   "Carrier_37_SpareSafetyOutput(3_4)" AT %I2215.4 : Bool;   // SPARE SAFETY OUTPUT
   "Carrier_37_SpareSafetyOutput(3_5)" AT %I2215.5 : Bool;   // SPARE SAFETY OUTPUT
   "Carrier_37_SpareSafetyOutput(3_6)" AT %I2215.6 : Bool;   // SPARE SAFETY OUTPUT
   "Carrier_37_SpareSafetyOutput(3_7)" AT %I2215.7 : Bool;   // SPARE SAFETY OUTPUT
   "Carrier_37_Slot4_Input" AT %IW2216 : Word;   // SLOT 4 INPUT WORD
   "Carrier_37_480VPowerOn_MDCB1" AT %I2216.0 : Bool;   // 480 VAC POWER ON MDCB 1
   "Carrier_37_SpareInput(4_1)" AT %I2216.1 : Bool;   // SPARE INPUT
   "Carrier_37_SpareInput(4_2)" AT %I2216.2 : Bool;   // SPARE INPUT
   "Carrier_37_SitopSelectStatus" AT %I2216.3 : Bool;   // SITOP SELECT STATUS
   "Carrier_37_DCsupplyOnPSCB2" AT %I2216.4 : Bool;   // DC SUPPLY ON PSCB 2
   "Carrier_37_SpareInput(4_5)" AT %I2216.5 : Bool;   // SPARE INPUT
   "Carrier_37_SpareInput(4_6)" AT %I2216.6 : Bool;   // SPARE INPUT
   "Carrier_37_SpareInput(4_7)" AT %I2216.7 : Bool;   // SPARE INPUT
   "Carrier_37_PB1_ProdHoldLH" AT %I2217.0 : Bool;   // PB 1 PRODUCTION HOLD LH
   "Carrier_37_PB2_ResetLH" AT %I2217.1 : Bool;   // PB 2 RESET LH
   "Carrier_37_PB3_ProdHoldRH" AT %I2217.2 : Bool;   // PB 3 PRODUCTION HOLD RH
   "Carrier_37_PB4_ResetRH" AT %I2217.3 : Bool;   // PB 4 RESET RH
   "Carrier_37_SpareInput(4_14)" AT %I2217.4 : Bool;   // SPARE INPUT
   "Carrier_37_SpareInput(4_15)" AT %I2217.5 : Bool;   // SPARE INPUT
   "Carrier_37_SpareInput(4_16)" AT %I2217.6 : Bool;   // SPARE INPUT
   "Carrier_37_SpareInput(4_17)" AT %I2217.7 : Bool;   // SPARE INPUT
   "Carrier_37_Slot5_Output" AT %IW2218 : Word;   // SLOT 5 OUTPUT WORD
   "Carrier_37_IRD400_HMI_24VDC_ENABLE" AT %I2218.0 : Bool;   // IRD 400 PANEL HMI 24V DC POWER
   "Carrier_37_FaultLight_LH" AT %I2218.1 : Bool;   // FAULT LIGHT LH
   "Carrier_37_RunLight_LH" AT %I2218.2 : Bool;   // RUN LIGHT LH
   "Carrier_37_FaultLight_RH" AT %I2218.3 : Bool;   // FAULT LIGHT RH
   "Carrier_37_RunLight_RH" AT %I2218.4 : Bool;   // RUN LIGHT RH
   "Carrier_37_SpareOutput(5_5)" AT %I2218.5 : Bool;   // SPARE OUTPUT
   "Carrier_37_SpareOutput(5_6)" AT %I2218.6 : Bool;   // SPARE OUTPUT
   "Carrier_37_SpareOutput(5_7)" AT %I2218.7 : Bool;   // SPARE OUTPUT
   "Carrier_37_ActualSpeed" AT %IW2220 : Word;   // ACTUAL SPEED
   "Carrier_37_CarrierDriveAlarm" AT %IW2222 : Word;   // CARRIER DRIVE ALARM
   "Carrier_37_CarrierDriveWarning" AT %IW2224 : Word;   // CARRIER DRIVE WARNING
   "Carrier_38_Status" AT %IW2250 : Word;   // CARRIER STATUS WORD
   "Carrier_38_Status.0" AT %I2250.0 : Bool;   // HEARTBEAT
   "Carrier_38_Status.1" AT %I2250.1 : Bool;   // MANUAL
   "Carrier_38_Status.2" AT %I2250.2 : Bool;   // IN_AUTO
   "Carrier_38_Status.3" AT %I2250.3 : Bool;   // POSITIONING_COMPLETE
   "Carrier_38_Status.4" AT %I2250.4 : Bool;   // PRODUCTION HOLD
   "Carrier_38_Status.5" AT %I2250.5 : Bool;   // CARRIER MOVING FORWARD
   "Carrier_38_Status.6" AT %I2250.6 : Bool;   // CARRIER MOVING REVERSE
   "Carrier_38_Status.7" AT %I2250.7 : Bool;   // CARRIER FAULT
   "Carrier_38_Status.8" AT %I2251.0 : Bool;   // CRASH DETECT TRIPPED
   "Carrier_38_Status.9" AT %I2251.1 : Bool;
   "Carrier_38_Status.10" AT %I2251.2 : Bool;
   "Carrier_38_Status.11" AT %I2251.3 : Bool;
   "Carrier_38_Status.12" AT %I2251.4 : Bool;
   "Carrier_38_Status.13" AT %I2251.5 : Bool;
   "Carrier_38_Status.14" AT %I2251.6 : Bool;
   "Carrier_38_Status.15" AT %I2251.7 : Bool;
   "Carrier_38_SDCFaultCode" AT %IW2252 : Word;   // SDC FAULT CODE
   "Carrier_38_CarrierPosition" AT %ID2254 : DWord;   // CARRIER POSITION
   "Carrier_38_CarrierNumber" AT %IW2258 : Word;   // CARRIER NUMBER
   "Carrier_38_G120DControlWord" AT %IW2260 : Word;   // G120D_STW1_CONTROL
   "Carrier_38_G120DControlWord.0" AT %I2260.0 : Bool;   // Bit_00_ON
   "Carrier_38_G120DControlWord.1" AT %I2260.1 : Bool;   // Bit_01_AUS2_INH
   "Carrier_38_G120DControlWord.2" AT %I2260.2 : Bool;   // Bit_02_AUS3_STOP
   "Carrier_38_G120DControlWord.3" AT %I2260.3 : Bool;   // Bit_03_EN
   "Carrier_38_G120DControlWord.4" AT %I2260.4 : Bool;   // Bit_04_EN_RAMP
   "Carrier_38_G120DControlWord.5" AT %I2260.5 : Bool;   // Bit_05_START_RAMP
   "Carrier_38_G120DControlWord.6" AT %I2260.6 : Bool;   // Bit_06_SETPOINT
   "Carrier_38_G120DControlWord.7" AT %I2260.7 : Bool;   // Bit_07_RESET
   "Carrier_38_G120DControlWord.8" AT %I2261.0 : Bool;   // Bit_08_JOG_R
   "Carrier_38_G120DControlWord.9" AT %I2261.1 : Bool;   // Bit_09_JOG_L
   "Carrier_38_G120DControlWord.10" AT %I2261.2 : Bool;   // Bit_10_CONTR_PLC
   "Carrier_38_G120DControlWord.11" AT %I2261.3 : Bool;   // Bit_11_REVERSE
   "Carrier_38_G120DControlWord.12" AT %I2261.4 : Bool;   // Bit_12_BRAKE_RELEASE
   "Carrier_38_G120DControlWord.13" AT %I2261.5 : Bool;   // Bit_13_DDS
   "Carrier_38_G120DControlWord.14" AT %I2261.6 : Bool;   // Bit_14_DO0
   "Carrier_38_G120DControlWord.15" AT %I2261.7 : Bool;   // Bit_15_DO1
   "Carrier_38_G120DStatusWord" AT %IW2262 : Word;   // G120D_ZSW1_STATUS
   "Carrier_38_G120DStatusWord.0" AT %I2262.0 : Bool;   // Bit_00_READY_RUN
   "Carrier_38_G120DStatusWord.1" AT %I2262.1 : Bool;   // Bit_01_READY_ON
   "Carrier_38_G120DStatusWord.2" AT %I2262.2 : Bool;   // Bit_02_ENABLE
   "Carrier_38_G120DStatusWord.3" AT %I2262.3 : Bool;   // Bit_03_FAULT
   "Carrier_38_G120DStatusWord.4" AT %I2262.4 : Bool;   // Bit_04_OFF2
   "Carrier_38_G120DStatusWord.5" AT %I2262.5 : Bool;   // Bit_05_OFF3
   "Carrier_38_G120DStatusWord.6" AT %I2262.6 : Bool;   // Bit_06_LOCK_OUT
   "Carrier_38_G120DStatusWord.7" AT %I2262.7 : Bool;   // Bit_07_WARN
   "Carrier_38_G120DStatusWord.8" AT %I2263.0 : Bool;   // Bit_08_NO_DEVIATION
   "Carrier_38_G120DStatusWord.9" AT %I2263.1 : Bool;   // Bit_09_CONTR_PLC
   "Carrier_38_G120DStatusWord.10" AT %I2263.2 : Bool;   // Bit_10_F_MAX
   "Carrier_38_G120DStatusWord.11" AT %I2263.3 : Bool;   // Bit_11_LIMIT_REACHED
   "Carrier_38_G120DStatusWord.12" AT %I2263.4 : Bool;   // Bit_12_BRAKE_OPEN
   "Carrier_38_G120DStatusWord.13" AT %I2263.5 : Bool;   // Bit_13_NO_OVERTEMP
   "Carrier_38_G120DStatusWord.14" AT %I2263.6 : Bool;   // Bit_14_CW_CCW
   "Carrier_38_G120DStatusWord.15" AT %I2263.7 : Bool;   // Bit_15_OVERL
   "Carrier_38_Slot2_Input" AT %IW2264 : Word;   // SLOT 2 INPUT WORD
   "Carrier_38_CrashDetectSW" AT %I2264.0 : Bool;   // CRASH DETECT SW
   "Carrier_38_SpareSafetyInput(2_1)" AT %I2264.1 : Bool;   // SPARE SAFETY INPUT
   "Carrier_38_SpareSafetyInput(2_2)" AT %I2264.2 : Bool;   // SPARE SAFETY INPUT
   "Carrier_38_SpareSafetyInput(2_3)" AT %I2264.3 : Bool;   // SPARE SAFETY INPUT
   "Carrier_38_SpareSafetyInput(2_4)" AT %I2264.4 : Bool;   // SPARE SAFETY INPUT
   "Carrier_38_SpareSafetyInput(2_5)" AT %I2264.5 : Bool;   // SPARE SAFETY INPUT
   "Carrier_38_SpareSafetyInput(2_6)" AT %I2264.6 : Bool;   // SPARE SAFETY INPUT
   "Carrier_38_SpareSafetyInput(2_7)" AT %I2264.7 : Bool;   // SPARE SAFETY INPUT
   "Carrier_38_Slot3_SafetyOutput" AT %IW2265 : Word;   // SLOT 3 SAFETY OUTPUT WORD
   "Carrier_38_Crash_Detect_OK" AT %I2265.0 : Bool;   // CARRIER CRASH DETECT
   "Carrier_38_SpareSafetyOutput(3_1)" AT %I2265.1 : Bool;   // SPARE SAFETY OUTPUT
   "Carrier_38_SpareSafetyOutput(3_2)" AT %I2265.2 : Bool;   // SPARE SAFETY OUTPUT
   "Carrier_38_SpareSafetyOutput(3_3)" AT %I2265.3 : Bool;   // SPARE SAFETY OUTPUT
   "Carrier_38_SpareSafetyOutput(3_4)" AT %I2265.4 : Bool;   // SPARE SAFETY OUTPUT
   "Carrier_38_SpareSafetyOutput(3_5)" AT %I2265.5 : Bool;   // SPARE SAFETY OUTPUT
   "Carrier_38_SpareSafetyOutput(3_6)" AT %I2265.6 : Bool;   // SPARE SAFETY OUTPUT
   "Carrier_38_SpareSafetyOutput(3_7)" AT %I2265.7 : Bool;   // SPARE SAFETY OUTPUT
   "Carrier_38_Slot4_Input" AT %IW2266 : Word;   // SLOT 4 INPUT WORD
   "Carrier_38_480VPowerOn_MDCB1" AT %I2266.0 : Bool;   // 480 VAC POWER ON MDCB 1
   "Carrier_38_SpareInput(4_1)" AT %I2266.1 : Bool;   // SPARE INPUT
   "Carrier_38_SpareInput(4_2)" AT %I2266.2 : Bool;   // SPARE INPUT
   "Carrier_38_SitopSelectStatus" AT %I2266.3 : Bool;   // SITOP SELECT STATUS
   "Carrier_38_DCsupplyOnPSCB2" AT %I2266.4 : Bool;   // DC SUPPLY ON PSCB 2
   "Carrier_38_SpareInput(4_5)" AT %I2266.5 : Bool;   // SPARE INPUT
   "Carrier_38_SpareInput(4_6)" AT %I2266.6 : Bool;   // SPARE INPUT
   "Carrier_38_SpareInput(4_7)" AT %I2266.7 : Bool;   // SPARE INPUT
   "Carrier_38_PB1_ProdHoldLH" AT %I2267.0 : Bool;   // PB 1 PRODUCTION HOLD LH
   "Carrier_38_PB2_ResetLH" AT %I2267.1 : Bool;   // PB 2 RESET LH
   "Carrier_38_PB3_ProdHoldRH" AT %I2267.2 : Bool;   // PB 3 PRODUCTION HOLD RH
   "Carrier_38_PB4_ResetRH" AT %I2267.3 : Bool;   // PB 4 RESET RH
   "Carrier_38_SpareInput(4_14)" AT %I2267.4 : Bool;   // SPARE INPUT
   "Carrier_38_SpareInput(4_15)" AT %I2267.5 : Bool;   // SPARE INPUT
   "Carrier_38_SpareInput(4_16)" AT %I2267.6 : Bool;   // SPARE INPUT
   "Carrier_38_SpareInput(4_17)" AT %I2267.7 : Bool;   // SPARE INPUT
   "Carrier_38_Slot5_Output" AT %IW2268 : Word;   // SLOT 5 OUTPUT WORD
   "Carrier_38_IRD400_HMI_24VDC_ENABLE" AT %I2268.0 : Bool;   // IRD 400 PANEL HMI 24V DC POWER
   "Carrier_38_FaultLight_LH" AT %I2268.1 : Bool;   // FAULT LIGHT LH
   "Carrier_38_RunLight_LH" AT %I2268.2 : Bool;   // RUN LIGHT LH
   "Carrier_38_FaultLight_RH" AT %I2268.3 : Bool;   // FAULT LIGHT RH
   "Carrier_38_RunLight_RH" AT %I2268.4 : Bool;   // RUN LIGHT RH
   "Carrier_38_SpareOutput(5_5)" AT %I2268.5 : Bool;   // SPARE OUTPUT
   "Carrier_38_SpareOutput(5_6)" AT %I2268.6 : Bool;   // SPARE OUTPUT
   "Carrier_38_SpareOutput(5_7)" AT %I2268.7 : Bool;   // SPARE OUTPUT
   "Carrier_38_ActualSpeed" AT %IW2270 : Word;   // ACTUAL SPEED
   "Carrier_38_CarrierDriveAlarm" AT %IW2272 : Word;   // CARRIER DRIVE ALARM
   "Carrier_38_CarrierDriveWarning" AT %IW2274 : Word;   // CARRIER DRIVE WARNING
   "Carrier_39_Status" AT %IW2300 : Word;   // CARRIER STATUS WORD
   "Carrier_39_Status.0" AT %I2300.0 : Bool;   // HEARTBEAT
   "Carrier_39_Status.1" AT %I2300.1 : Bool;   // MANUAL
   "Carrier_39_Status.2" AT %I2300.2 : Bool;   // IN_AUTO
   "Carrier_39_Status.3" AT %I2300.3 : Bool;   // POSITIONING_COMPLETE
   "Carrier_39_Status.4" AT %I2300.4 : Bool;   // PRODUCTION HOLD
   "Carrier_39_Status.5" AT %I2300.5 : Bool;   // CARRIER MOVING FORWARD
   "Carrier_39_Status.6" AT %I2300.6 : Bool;   // CARRIER MOVING REVERSE
   "Carrier_39_Status.7" AT %I2300.7 : Bool;   // CARRIER FAULT
   "Carrier_39_Status.8" AT %I2301.0 : Bool;   // CRASH DETECT TRIPPED
   "Carrier_39_Status.9" AT %I2301.1 : Bool;
   "Carrier_39_Status.10" AT %I2301.2 : Bool;
   "Carrier_39_Status.11" AT %I2301.3 : Bool;
   "Carrier_39_Status.12" AT %I2301.4 : Bool;
   "Carrier_39_Status.13" AT %I2301.5 : Bool;
   "Carrier_39_Status.14" AT %I2301.6 : Bool;
   "Carrier_39_Status.15" AT %I2301.7 : Bool;
   "Carrier_39_SDCFaultCode" AT %IW2302 : Word;   // SDC FAULT CODE
   "Carrier_39_CarrierPosition" AT %ID2304 : DWord;   // CARRIER POSITION
   "Carrier_39_CarrierNumber" AT %IW2308 : Word;   // CARRIER NUMBER
   "Carrier_39_G120DControlWord" AT %IW2310 : Word;   // G120D_STW1_CONTROL
   "Carrier_39_G120DControlWord.0" AT %I2310.0 : Bool;   // Bit_00_ON
   "Carrier_39_G120DControlWord.1" AT %I2310.1 : Bool;   // Bit_01_AUS2_INH
   "Carrier_39_G120DControlWord.2" AT %I2310.2 : Bool;   // Bit_02_AUS3_STOP
   "Carrier_39_G120DControlWord.3" AT %I2310.3 : Bool;   // Bit_03_EN
   "Carrier_39_G120DControlWord.4" AT %I2310.4 : Bool;   // Bit_04_EN_RAMP
   "Carrier_39_G120DControlWord.5" AT %I2310.5 : Bool;   // Bit_05_START_RAMP
   "Carrier_39_G120DControlWord.6" AT %I2310.6 : Bool;   // Bit_06_SETPOINT
   "Carrier_39_G120DControlWord.7" AT %I2310.7 : Bool;   // Bit_07_RESET
   "Carrier_39_G120DControlWord.8" AT %I2311.0 : Bool;   // Bit_08_JOG_R
   "Carrier_39_G120DControlWord.9" AT %I2311.1 : Bool;   // Bit_09_JOG_L
   "Carrier_39_G120DControlWord.10" AT %I2311.2 : Bool;   // Bit_10_CONTR_PLC
   "Carrier_39_G120DControlWord.11" AT %I2311.3 : Bool;   // Bit_11_REVERSE
   "Carrier_39_G120DControlWord.12" AT %I2311.4 : Bool;   // Bit_12_BRAKE_RELEASE
   "Carrier_39_G120DControlWord.13" AT %I2311.5 : Bool;   // Bit_13_DDS
   "Carrier_39_G120DControlWord.14" AT %I2311.6 : Bool;   // Bit_14_DO0
   "Carrier_39_G120DControlWord.15" AT %I2311.7 : Bool;   // Bit_15_DO1
   "Carrier_39_G120DStatusWord" AT %IW2312 : Word;   // G120D_ZSW1_STATUS
   "Carrier_39_G120DStatusWord.0" AT %I2312.0 : Bool;   // Bit_00_READY_RUN
   "Carrier_39_G120DStatusWord.1" AT %I2312.1 : Bool;   // Bit_01_READY_ON
   "Carrier_39_G120DStatusWord.2" AT %I2312.2 : Bool;   // Bit_02_ENABLE
   "Carrier_39_G120DStatusWord.3" AT %I2312.3 : Bool;   // Bit_03_FAULT
   "Carrier_39_G120DStatusWord.4" AT %I2312.4 : Bool;   // Bit_04_OFF2
   "Carrier_39_G120DStatusWord.5" AT %I2312.5 : Bool;   // Bit_05_OFF3
   "Carrier_39_G120DStatusWord.6" AT %I2312.6 : Bool;   // Bit_06_LOCK_OUT
   "Carrier_39_G120DStatusWord.7" AT %I2312.7 : Bool;   // Bit_07_WARN
   "Carrier_39_G120DStatusWord.8" AT %I2313.0 : Bool;   // Bit_08_NO_DEVIATION
   "Carrier_39_G120DStatusWord.9" AT %I2313.1 : Bool;   // Bit_09_CONTR_PLC
   "Carrier_39_G120DStatusWord.10" AT %I2313.2 : Bool;   // Bit_10_F_MAX
   "Carrier_39_G120DStatusWord.11" AT %I2313.3 : Bool;   // Bit_11_LIMIT_REACHED
   "Carrier_39_G120DStatusWord.12" AT %I2313.4 : Bool;   // Bit_12_BRAKE_OPEN
   "Carrier_39_G120DStatusWord.13" AT %I2313.5 : Bool;   // Bit_13_NO_OVERTEMP
   "Carrier_39_G120DStatusWord.14" AT %I2313.6 : Bool;   // Bit_14_CW_CCW
   "Carrier_39_G120DStatusWord.15" AT %I2313.7 : Bool;   // Bit_15_OVERL
   "Carrier_39_Slot2_Input" AT %IW2314 : Word;   // SLOT 2 INPUT WORD
   "Carrier_39_CrashDetectSW" AT %I2314.0 : Bool;   // CRASH DETECT SW
   "Carrier_39_SpareSafetyInput(2_1)" AT %I2314.1 : Bool;   // SPARE SAFETY INPUT
   "Carrier_39_SpareSafetyInput(2_2)" AT %I2314.2 : Bool;   // SPARE SAFETY INPUT
   "Carrier_39_SpareSafetyInput(2_3)" AT %I2314.3 : Bool;   // SPARE SAFETY INPUT
   "Carrier_39_SpareSafetyInput(2_4)" AT %I2314.4 : Bool;   // SPARE SAFETY INPUT
   "Carrier_39_SpareSafetyInput(2_5)" AT %I2314.5 : Bool;   // SPARE SAFETY INPUT
   "Carrier_39_SpareSafetyInput(2_6)" AT %I2314.6 : Bool;   // SPARE SAFETY INPUT
   "Carrier_39_SpareSafetyInput(2_7)" AT %I2314.7 : Bool;   // SPARE SAFETY INPUT
   "Carrier_39_Slot3_SafetyOutput" AT %IW2315 : Word;   // SLOT 3 SAFETY OUTPUT WORD
   "Carrier_39_Crash_Detect_OK" AT %I2315.0 : Bool;   // CARRIER CRASH DETECT
   "Carrier_39_SpareSafetyOutput(3_1)" AT %I2315.1 : Bool;   // SPARE SAFETY OUTPUT
   "Carrier_39_SpareSafetyOutput(3_2)" AT %I2315.2 : Bool;   // SPARE SAFETY OUTPUT
   "Carrier_39_SpareSafetyOutput(3_3)" AT %I2315.3 : Bool;   // SPARE SAFETY OUTPUT
   "Carrier_39_SpareSafetyOutput(3_4)" AT %I2315.4 : Bool;   // SPARE SAFETY OUTPUT
   "Carrier_39_SpareSafetyOutput(3_5)" AT %I2315.5 : Bool;   // SPARE SAFETY OUTPUT
   "Carrier_39_SpareSafetyOutput(3_6)" AT %I2315.6 : Bool;   // SPARE SAFETY OUTPUT
   "Carrier_39_SpareSafetyOutput(3_7)" AT %I2315.7 : Bool;   // SPARE SAFETY OUTPUT
   "Carrier_39_Slot4_Input" AT %IW2316 : Word;   // SLOT 4 INPUT WORD
   "Carrier_39_480VPowerOn_MDCB1" AT %I2316.0 : Bool;   // 480 VAC POWER ON MDCB 1
   "Carrier_39_SpareInput(4_1)" AT %I2316.1 : Bool;   // SPARE INPUT
   "Carrier_39_SpareInput(4_2)" AT %I2316.2 : Bool;   // SPARE INPUT
   "Carrier_39_SitopSelectStatus" AT %I2316.3 : Bool;   // SITOP SELECT STATUS
   "Carrier_39_DCsupplyOnPSCB2" AT %I2316.4 : Bool;   // DC SUPPLY ON PSCB 2
   "Carrier_39_SpareInput(4_5)" AT %I2316.5 : Bool;   // SPARE INPUT
   "Carrier_39_SpareInput(4_6)" AT %I2316.6 : Bool;   // SPARE INPUT
   "Carrier_39_SpareInput(4_7)" AT %I2316.7 : Bool;   // SPARE INPUT
   "Carrier_39_PB1_ProdHoldLH" AT %I2317.0 : Bool;   // PB 1 PRODUCTION HOLD LH
   "Carrier_39_PB2_ResetLH" AT %I2317.1 : Bool;   // PB 2 RESET LH
   "Carrier_39_PB3_ProdHoldRH" AT %I2317.2 : Bool;   // PB 3 PRODUCTION HOLD RH
   "Carrier_39_PB4_ResetRH" AT %I2317.3 : Bool;   // PB 4 RESET RH
   "Carrier_39_SpareInput(4_14)" AT %I2317.4 : Bool;   // SPARE INPUT
   "Carrier_39_SpareInput(4_15)" AT %I2317.5 : Bool;   // SPARE INPUT
   "Carrier_39_SpareInput(4_16)" AT %I2317.6 : Bool;   // SPARE INPUT
   "Carrier_39_SpareInput(4_17)" AT %I2317.7 : Bool;   // SPARE INPUT
   "Carrier_39_Slot5_Output" AT %IW2318 : Word;   // SLOT 5 OUTPUT WORD
   "Carrier_39_IRD400_HMI_24VDC_ENABLE" AT %I2318.0 : Bool;   // IRD 400 PANEL HMI 24V DC POWER
   "Carrier_39_FaultLight_LH" AT %I2318.1 : Bool;   // FAULT LIGHT LH
   "Carrier_39_RunLight_LH" AT %I2318.2 : Bool;   // RUN LIGHT LH
   "Carrier_39_FaultLight_RH" AT %I2318.3 : Bool;   // FAULT LIGHT RH
   "Carrier_39_RunLight_RH" AT %I2318.4 : Bool;   // RUN LIGHT RH
   "Carrier_39_SpareOutput(5_5)" AT %I2318.5 : Bool;   // SPARE OUTPUT
   "Carrier_39_SpareOutput(5_6)" AT %I2318.6 : Bool;   // SPARE OUTPUT
   "Carrier_39_SpareOutput(5_7)" AT %I2318.7 : Bool;   // SPARE OUTPUT
   "Carrier_39_ActualSpeed" AT %IW2320 : Word;   // ACTUAL SPEED
   "Carrier_39_CarrierDriveAlarm" AT %IW2322 : Word;   // CARRIER DRIVE ALARM
   "Carrier_39_CarrierDriveWarning" AT %IW2324 : Word;   // CARRIER DRIVE WARNING
   "Carrier_40_Status" AT %IW2350 : Word;   // CARRIER STATUS WORD
   "Carrier_40_Status.0" AT %I2350.0 : Bool;   // HEARTBEAT
   "Carrier_40_Status.1" AT %I2350.1 : Bool;   // MANUAL
   "Carrier_40_Status.2" AT %I2350.2 : Bool;   // IN_AUTO
   "Carrier_40_Status.3" AT %I2350.3 : Bool;   // POSITIONING_COMPLETE
   "Carrier_40_Status.4" AT %I2350.4 : Bool;   // PRODUCTION HOLD
   "Carrier_40_Status.5" AT %I2350.5 : Bool;   // CARRIER MOVING FORWARD
   "Carrier_40_Status.6" AT %I2350.6 : Bool;   // CARRIER MOVING REVERSE
   "Carrier_40_Status.7" AT %I2350.7 : Bool;   // CARRIER FAULT
   "Carrier_40_Status.8" AT %I2351.0 : Bool;   // CRASH DETECT TRIPPED
   "Carrier_40_Status.9" AT %I2351.1 : Bool;
   "Carrier_40_Status.10" AT %I2351.2 : Bool;
   "Carrier_40_Status.11" AT %I2351.3 : Bool;
   "Carrier_40_Status.12" AT %I2351.4 : Bool;
   "Carrier_40_Status.13" AT %I2351.5 : Bool;
   "Carrier_40_Status.14" AT %I2351.6 : Bool;
   "Carrier_40_Status.15" AT %I2351.7 : Bool;
   "Carrier_40_SDCFaultCode" AT %IW2352 : Word;   // SDC FAULT CODE
   "Carrier_40_CarrierPosition" AT %ID2354 : DWord;   // CARRIER POSITION
   "Carrier_40_CarrierNumber" AT %IW2358 : Word;   // CARRIER NUMBER
   "Carrier_40_G120DControlWord" AT %IW2360 : Word;   // G120D_STW1_CONTROL
   "Carrier_40_G120DControlWord.0" AT %I2360.0 : Bool;   // Bit_00_ON
   "Carrier_40_G120DControlWord.1" AT %I2360.1 : Bool;   // Bit_01_AUS2_INH
   "Carrier_40_G120DControlWord.2" AT %I2360.2 : Bool;   // Bit_02_AUS3_STOP
   "Carrier_40_G120DControlWord.3" AT %I2360.3 : Bool;   // Bit_03_EN
   "Carrier_40_G120DControlWord.4" AT %I2360.4 : Bool;   // Bit_04_EN_RAMP
   "Carrier_40_G120DControlWord.5" AT %I2360.5 : Bool;   // Bit_05_START_RAMP
   "Carrier_40_G120DControlWord.6" AT %I2360.6 : Bool;   // Bit_06_SETPOINT
   "Carrier_40_G120DControlWord.7" AT %I2360.7 : Bool;   // Bit_07_RESET
   "Carrier_40_G120DControlWord.8" AT %I2361.0 : Bool;   // Bit_08_JOG_R
   "Carrier_40_G120DControlWord.9" AT %I2361.1 : Bool;   // Bit_09_JOG_L
   "Carrier_40_G120DControlWord.10" AT %I2361.2 : Bool;   // Bit_10_CONTR_PLC
   "Carrier_40_G120DControlWord.11" AT %I2361.3 : Bool;   // Bit_11_REVERSE
   "Carrier_40_G120DControlWord.12" AT %I2361.4 : Bool;   // Bit_12_BRAKE_RELEASE
   "Carrier_40_G120DControlWord.13" AT %I2361.5 : Bool;   // Bit_13_DDS
   "Carrier_40_G120DControlWord.14" AT %I2361.6 : Bool;   // Bit_14_DO0
   "Carrier_40_G120DControlWord.15" AT %I2361.7 : Bool;   // Bit_15_DO1
   "Carrier_40_G120DStatusWord" AT %IW2362 : Word;   // G120D_ZSW1_STATUS
   "Carrier_40_G120DStatusWord.0" AT %I2362.0 : Bool;   // Bit_00_READY_RUN
   "Carrier_40_G120DStatusWord.1" AT %I2362.1 : Bool;   // Bit_01_READY_ON
   "Carrier_40_G120DStatusWord.2" AT %I2362.2 : Bool;   // Bit_02_ENABLE
   "Carrier_40_G120DStatusWord.3" AT %I2362.3 : Bool;   // Bit_03_FAULT
   "Carrier_40_G120DStatusWord.4" AT %I2362.4 : Bool;   // Bit_04_OFF2
   "Carrier_40_G120DStatusWord.5" AT %I2362.5 : Bool;   // Bit_05_OFF3
   "Carrier_40_G120DStatusWord.6" AT %I2362.6 : Bool;   // Bit_06_LOCK_OUT
   "Carrier_40_G120DStatusWord.7" AT %I2362.7 : Bool;   // Bit_07_WARN
   "Carrier_40_G120DStatusWord.8" AT %I2363.0 : Bool;   // Bit_08_NO_DEVIATION
   "Carrier_40_G120DStatusWord.9" AT %I2363.1 : Bool;   // Bit_09_CONTR_PLC
   "Carrier_40_G120DStatusWord.10" AT %I2363.2 : Bool;   // Bit_10_F_MAX
   "Carrier_40_G120DStatusWord.11" AT %I2363.3 : Bool;   // Bit_11_LIMIT_REACHED
   "Carrier_40_G120DStatusWord.12" AT %I2363.4 : Bool;   // Bit_12_BRAKE_OPEN
   "Carrier_40_G120DStatusWord.13" AT %I2363.5 : Bool;   // Bit_13_NO_OVERTEMP
   "Carrier_40_G120DStatusWord.14" AT %I2363.6 : Bool;   // Bit_14_CW_CCW
   "Carrier_40_G120DStatusWord.15" AT %I2363.7 : Bool;   // Bit_15_OVERL
   "Carrier_40_Slot2_Input" AT %IW2364 : Word;   // SLOT 2 INPUT WORD
   "Carrier_40_CrashDetectSW" AT %I2364.0 : Bool;   // CRASH DETECT SW
   "Carrier_40_SpareSafetyInput(2_1)" AT %I2364.1 : Bool;   // SPARE SAFETY INPUT
   "Carrier_40_SpareSafetyInput(2_2)" AT %I2364.2 : Bool;   // SPARE SAFETY INPUT
   "Carrier_40_SpareSafetyInput(2_3)" AT %I2364.3 : Bool;   // SPARE SAFETY INPUT
   "Carrier_40_SpareSafetyInput(2_4)" AT %I2364.4 : Bool;   // SPARE SAFETY INPUT
   "Carrier_40_SpareSafetyInput(2_5)" AT %I2364.5 : Bool;   // SPARE SAFETY INPUT
   "Carrier_40_SpareSafetyInput(2_6)" AT %I2364.6 : Bool;   // SPARE SAFETY INPUT
   "Carrier_40_SpareSafetyInput(2_7)" AT %I2364.7 : Bool;   // SPARE SAFETY INPUT
   "Carrier_40_Slot3_SafetyOutput" AT %IW2365 : Word;   // SLOT 3 SAFETY OUTPUT WORD
   "Carrier_40_Crash_Detect_OK" AT %I2365.0 : Bool;   // CARRIER CRASH DETECT
   "Carrier_40_SpareSafetyOutput(3_1)" AT %I2365.1 : Bool;   // SPARE SAFETY OUTPUT
   "Carrier_40_SpareSafetyOutput(3_2)" AT %I2365.2 : Bool;   // SPARE SAFETY OUTPUT
   "Carrier_40_SpareSafetyOutput(3_3)" AT %I2365.3 : Bool;   // SPARE SAFETY OUTPUT
   "Carrier_40_SpareSafetyOutput(3_4)" AT %I2365.4 : Bool;   // SPARE SAFETY OUTPUT
   "Carrier_40_SpareSafetyOutput(3_5)" AT %I2365.5 : Bool;   // SPARE SAFETY OUTPUT
   "Carrier_40_SpareSafetyOutput(3_6)" AT %I2365.6 : Bool;   // SPARE SAFETY OUTPUT
   "Carrier_40_SpareSafetyOutput(3_7)" AT %I2365.7 : Bool;   // SPARE SAFETY OUTPUT
   "Carrier_40_Slot4_Input" AT %IW2366 : Word;   // SLOT 4 INPUT WORD
   "Carrier_40_480VPowerOn_MDCB1" AT %I2366.0 : Bool;   // 480 VAC POWER ON MDCB 1
   "Carrier_40_SpareInput(4_1)" AT %I2366.1 : Bool;   // SPARE INPUT
   "Carrier_40_SpareInput(4_2)" AT %I2366.2 : Bool;   // SPARE INPUT
   "Carrier_40_SitopSelectStatus" AT %I2366.3 : Bool;   // SITOP SELECT STATUS
   "Carrier_40_DCsupplyOnPSCB2" AT %I2366.4 : Bool;   // DC SUPPLY ON PSCB 2
   "Carrier_40_SpareInput(4_5)" AT %I2366.5 : Bool;   // SPARE INPUT
   "Carrier_40_SpareInput(4_6)" AT %I2366.6 : Bool;   // SPARE INPUT
   "Carrier_40_SpareInput(4_7)" AT %I2366.7 : Bool;   // SPARE INPUT
   "Carrier_40_PB1_ProdHoldLH" AT %I2367.0 : Bool;   // PB 1 PRODUCTION HOLD LH
   "Carrier_40_PB2_ResetLH" AT %I2367.1 : Bool;   // PB 2 RESET LH
   "Carrier_40_PB3_ProdHoldRH" AT %I2367.2 : Bool;   // PB 3 PRODUCTION HOLD RH
   "Carrier_40_PB4_ResetRH" AT %I2367.3 : Bool;   // PB 4 RESET RH
   "Carrier_40_SpareInput(4_14)" AT %I2367.4 : Bool;   // SPARE INPUT
   "Carrier_40_SpareInput(4_15)" AT %I2367.5 : Bool;   // SPARE INPUT
   "Carrier_40_SpareInput(4_16)" AT %I2367.6 : Bool;   // SPARE INPUT
   "Carrier_40_SpareInput(4_17)" AT %I2367.7 : Bool;   // SPARE INPUT
   "Carrier_40_Slot5_Output" AT %IW2368 : Word;   // SLOT 5 OUTPUT WORD
   "Carrier_40_IRD400_HMI_24VDC_ENABLE" AT %I2368.0 : Bool;   // IRD 400 PANEL HMI 24V DC POWER
   "Carrier_40_FaultLight_LH" AT %I2368.1 : Bool;   // FAULT LIGHT LH
   "Carrier_40_RunLight_LH" AT %I2368.2 : Bool;   // RUN LIGHT LH
   "Carrier_40_FaultLight_RH" AT %I2368.3 : Bool;   // FAULT LIGHT RH
   "Carrier_40_RunLight_RH" AT %I2368.4 : Bool;   // RUN LIGHT RH
   "Carrier_40_SpareOutput(5_5)" AT %I2368.5 : Bool;   // SPARE OUTPUT
   "Carrier_40_SpareOutput(5_6)" AT %I2368.6 : Bool;   // SPARE OUTPUT
   "Carrier_40_SpareOutput(5_7)" AT %I2368.7 : Bool;   // SPARE OUTPUT
   "Carrier_40_ActualSpeed" AT %IW2370 : Word;   // ACTUAL SPEED
   "Carrier_40_CarrierDriveAlarm" AT %IW2372 : Word;   // CARRIER DRIVE ALARM
   "Carrier_40_CarrierDriveWarning" AT %IW2374 : Word;   // CARRIER DRIVE WARNING
   "Carrier_41_Status" AT %IW2400 : Word;   // CARRIER STATUS WORD
   "Carrier_41_Status.0" AT %I2400.0 : Bool;   // HEARTBEAT
   "Carrier_41_Status.1" AT %I2400.1 : Bool;   // MANUAL
   "Carrier_41_Status.2" AT %I2400.2 : Bool;   // IN_AUTO
   "Carrier_41_Status.3" AT %I2400.3 : Bool;   // POSITIONING_COMPLETE
   "Carrier_41_Status.4" AT %I2400.4 : Bool;   // PRODUCTION HOLD
   "Carrier_41_Status.5" AT %I2400.5 : Bool;   // CARRIER MOVING FORWARD
   "Carrier_41_Status.6" AT %I2400.6 : Bool;   // CARRIER MOVING REVERSE
   "Carrier_41_Status.7" AT %I2400.7 : Bool;   // CARRIER FAULT
   "Carrier_41_Status.8" AT %I2401.0 : Bool;   // CRASH DETECT TRIPPED
   "Carrier_41_Status.9" AT %I2401.1 : Bool;
   "Carrier_41_Status.10" AT %I2401.2 : Bool;
   "Carrier_41_Status.11" AT %I2401.3 : Bool;
   "Carrier_41_Status.12" AT %I2401.4 : Bool;
   "Carrier_41_Status.13" AT %I2401.5 : Bool;
   "Carrier_41_Status.14" AT %I2401.6 : Bool;
   "Carrier_41_Status.15" AT %I2401.7 : Bool;
   "Carrier_41_SDCFaultCode" AT %IW2402 : Word;   // SDC FAULT CODE
   "Carrier_41_CarrierPosition" AT %ID2404 : DWord;   // CARRIER POSITION
   "Carrier_41_CarrierNumber" AT %IW2408 : Word;   // CARRIER NUMBER
   "Carrier_41_G120DControlWord" AT %IW2410 : Word;   // G120D_STW1_CONTROL
   "Carrier_41_G120DControlWord.0" AT %I2410.0 : Bool;   // Bit_00_ON
   "Carrier_41_G120DControlWord.1" AT %I2410.1 : Bool;   // Bit_01_AUS2_INH
   "Carrier_41_G120DControlWord.2" AT %I2410.2 : Bool;   // Bit_02_AUS3_STOP
   "Carrier_41_G120DControlWord.3" AT %I2410.3 : Bool;   // Bit_03_EN
   "Carrier_41_G120DControlWord.4" AT %I2410.4 : Bool;   // Bit_04_EN_RAMP
   "Carrier_41_G120DControlWord.5" AT %I2410.5 : Bool;   // Bit_05_START_RAMP
   "Carrier_41_G120DControlWord.6" AT %I2410.6 : Bool;   // Bit_06_SETPOINT
   "Carrier_41_G120DControlWord.7" AT %I2410.7 : Bool;   // Bit_07_RESET
   "Carrier_41_G120DControlWord.8" AT %I2411.0 : Bool;   // Bit_08_JOG_R
   "Carrier_41_G120DControlWord.9" AT %I2411.1 : Bool;   // Bit_09_JOG_L
   "Carrier_41_G120DControlWord.10" AT %I2411.2 : Bool;   // Bit_10_CONTR_PLC
   "Carrier_41_G120DControlWord.11" AT %I2411.3 : Bool;   // Bit_11_REVERSE
   "Carrier_41_G120DControlWord.12" AT %I2411.4 : Bool;   // Bit_12_BRAKE_RELEASE
   "Carrier_41_G120DControlWord.13" AT %I2411.5 : Bool;   // Bit_13_DDS
   "Carrier_41_G120DControlWord.14" AT %I2411.6 : Bool;   // Bit_14_DO0
   "Carrier_41_G120DControlWord.15" AT %I2411.7 : Bool;   // Bit_15_DO1
   "Carrier_41_G120DStatusWord" AT %IW2412 : Word;   // G120D_ZSW1_STATUS
   "Carrier_41_G120DStatusWord.0" AT %I2412.0 : Bool;   // Bit_00_READY_RUN
   "Carrier_41_G120DStatusWord.1" AT %I2412.1 : Bool;   // Bit_01_READY_ON
   "Carrier_41_G120DStatusWord.2" AT %I2412.2 : Bool;   // Bit_02_ENABLE
   "Carrier_41_G120DStatusWord.3" AT %I2412.3 : Bool;   // Bit_03_FAULT
   "Carrier_41_G120DStatusWord.4" AT %I2412.4 : Bool;   // Bit_04_OFF2
   "Carrier_41_G120DStatusWord.5" AT %I2412.5 : Bool;   // Bit_05_OFF3
   "Carrier_41_G120DStatusWord.6" AT %I2412.6 : Bool;   // Bit_06_LOCK_OUT
   "Carrier_41_G120DStatusWord.7" AT %I2412.7 : Bool;   // Bit_07_WARN
   "Carrier_41_G120DStatusWord.8" AT %I2413.0 : Bool;   // Bit_08_NO_DEVIATION
   "Carrier_41_G120DStatusWord.9" AT %I2413.1 : Bool;   // Bit_09_CONTR_PLC
   "Carrier_41_G120DStatusWord.10" AT %I2413.2 : Bool;   // Bit_10_F_MAX
   "Carrier_41_G120DStatusWord.11" AT %I2413.3 : Bool;   // Bit_11_LIMIT_REACHED
   "Carrier_41_G120DStatusWord.12" AT %I2413.4 : Bool;   // Bit_12_BRAKE_OPEN
   "Carrier_41_G120DStatusWord.13" AT %I2413.5 : Bool;   // Bit_13_NO_OVERTEMP
   "Carrier_41_G120DStatusWord.14" AT %I2413.6 : Bool;   // Bit_14_CW_CCW
   "Carrier_41_G120DStatusWord.15" AT %I2413.7 : Bool;   // Bit_15_OVERL
   "Carrier_41_Slot2_Input" AT %IW2414 : Word;   // SLOT 2 INPUT WORD
   "Carrier_41_CrashDetectSW" AT %I2414.0 : Bool;   // CRASH DETECT SW
   "Carrier_41_SpareSafetyInput(2_1)" AT %I2414.1 : Bool;   // SPARE SAFETY INPUT
   "Carrier_41_SpareSafetyInput(2_2)" AT %I2414.2 : Bool;   // SPARE SAFETY INPUT
   "Carrier_41_SpareSafetyInput(2_3)" AT %I2414.3 : Bool;   // SPARE SAFETY INPUT
   "Carrier_41_SpareSafetyInput(2_4)" AT %I2414.4 : Bool;   // SPARE SAFETY INPUT
   "Carrier_41_SpareSafetyInput(2_5)" AT %I2414.5 : Bool;   // SPARE SAFETY INPUT
   "Carrier_41_SpareSafetyInput(2_6)" AT %I2414.6 : Bool;   // SPARE SAFETY INPUT
   "Carrier_41_SpareSafetyInput(2_7)" AT %I2414.7 : Bool;   // SPARE SAFETY INPUT
   "Carrier_41_Slot3_SafetyOutput" AT %IW2415 : Word;   // SLOT 3 SAFETY OUTPUT WORD
   "Carrier_41_Crash_Detect_OK" AT %I2415.0 : Bool;   // CARRIER CRASH DETECT
   "Carrier_41_SpareSafetyOutput(3_1)" AT %I2415.1 : Bool;   // SPARE SAFETY OUTPUT
   "Carrier_41_SpareSafetyOutput(3_2)" AT %I2415.2 : Bool;   // SPARE SAFETY OUTPUT
   "Carrier_41_SpareSafetyOutput(3_3)" AT %I2415.3 : Bool;   // SPARE SAFETY OUTPUT
   "Carrier_41_SpareSafetyOutput(3_4)" AT %I2415.4 : Bool;   // SPARE SAFETY OUTPUT
   "Carrier_41_SpareSafetyOutput(3_5)" AT %I2415.5 : Bool;   // SPARE SAFETY OUTPUT
   "Carrier_41_SpareSafetyOutput(3_6)" AT %I2415.6 : Bool;   // SPARE SAFETY OUTPUT
   "Carrier_41_SpareSafetyOutput(3_7)" AT %I2415.7 : Bool;   // SPARE SAFETY OUTPUT
   "Carrier_41_Slot4_Input" AT %IW2416 : Word;   // SLOT 4 INPUT WORD
   "Carrier_41_480VPowerOn_MDCB1" AT %I2416.0 : Bool;   // 480 VAC POWER ON MDCB 1
   "Carrier_41_SpareInput(4_1)" AT %I2416.1 : Bool;   // SPARE INPUT
   "Carrier_41_SpareInput(4_2)" AT %I2416.2 : Bool;   // SPARE INPUT
   "Carrier_41_SitopSelectStatus" AT %I2416.3 : Bool;   // SITOP SELECT STATUS
   "Carrier_41_DCsupplyOnPSCB2" AT %I2416.4 : Bool;   // DC SUPPLY ON PSCB 2
   "Carrier_41_SpareInput(4_5)" AT %I2416.5 : Bool;   // SPARE INPUT
   "Carrier_41_SpareInput(4_6)" AT %I2416.6 : Bool;   // SPARE INPUT
   "Carrier_41_SpareInput(4_7)" AT %I2416.7 : Bool;   // SPARE INPUT
   "Carrier_41_PB1_ProdHoldLH" AT %I2417.0 : Bool;   // PB 1 PRODUCTION HOLD LH
   "Carrier_41_PB2_ResetLH" AT %I2417.1 : Bool;   // PB 2 RESET LH
   "Carrier_41_PB3_ProdHoldRH" AT %I2417.2 : Bool;   // PB 3 PRODUCTION HOLD RH
   "Carrier_41_PB4_ResetRH" AT %I2417.3 : Bool;   // PB 4 RESET RH
   "Carrier_41_SpareInput(4_14)" AT %I2417.4 : Bool;   // SPARE INPUT
   "Carrier_41_SpareInput(4_15)" AT %I2417.5 : Bool;   // SPARE INPUT
   "Carrier_41_SpareInput(4_16)" AT %I2417.6 : Bool;   // SPARE INPUT
   "Carrier_41_SpareInput(4_17)" AT %I2417.7 : Bool;   // SPARE INPUT
   "Carrier_41_Slot5_Output" AT %IW2418 : Word;   // SLOT 5 OUTPUT WORD
   "Carrier_41_IRD400_HMI_24VDC_ENABLE" AT %I2418.0 : Bool;   // IRD 400 PANEL HMI 24V DC POWER
   "Carrier_41_FaultLight_LH" AT %I2418.1 : Bool;   // FAULT LIGHT LH
   "Carrier_41_RunLight_LH" AT %I2418.2 : Bool;   // RUN LIGHT LH
   "Carrier_41_FaultLight_RH" AT %I2418.3 : Bool;   // FAULT LIGHT RH
   "Carrier_41_RunLight_RH" AT %I2418.4 : Bool;   // RUN LIGHT RH
   "Carrier_41_SpareOutput(5_5)" AT %I2418.5 : Bool;   // SPARE OUTPUT
   "Carrier_41_SpareOutput(5_6)" AT %I2418.6 : Bool;   // SPARE OUTPUT
   "Carrier_41_SpareOutput(5_7)" AT %I2418.7 : Bool;   // SPARE OUTPUT
   "Carrier_41_ActualSpeed" AT %IW2420 : Word;   // ACTUAL SPEED
   "Carrier_41_CarrierDriveAlarm" AT %IW2422 : Word;   // CARRIER DRIVE ALARM
   "Carrier_41_CarrierDriveWarning" AT %IW2424 : Word;   // CARRIER DRIVE WARNING
   "Carrier_42_Status" AT %IW2450 : Word;   // CARRIER STATUS WORD
   "Carrier_42_Status.0" AT %I2450.0 : Bool;   // HEARTBEAT
   "Carrier_42_Status.1" AT %I2450.1 : Bool;   // MANUAL
   "Carrier_42_Status.2" AT %I2450.2 : Bool;   // IN_AUTO
   "Carrier_42_Status.3" AT %I2450.3 : Bool;   // POSITIONING_COMPLETE
   "Carrier_42_Status.4" AT %I2450.4 : Bool;   // PRODUCTION HOLD
   "Carrier_42_Status.5" AT %I2450.5 : Bool;   // CARRIER MOVING FORWARD
   "Carrier_42_Status.6" AT %I2450.6 : Bool;   // CARRIER MOVING REVERSE
   "Carrier_42_Status.7" AT %I2450.7 : Bool;   // CARRIER FAULT
   "Carrier_42_Status.8" AT %I2451.0 : Bool;   // CRASH DETECT TRIPPED
   "Carrier_42_Status.9" AT %I2451.1 : Bool;
   "Carrier_42_Status.10" AT %I2451.2 : Bool;
   "Carrier_42_Status.11" AT %I2451.3 : Bool;
   "Carrier_42_Status.12" AT %I2451.4 : Bool;
   "Carrier_42_Status.13" AT %I2451.5 : Bool;
   "Carrier_42_Status.14" AT %I2451.6 : Bool;
   "Carrier_42_Status.15" AT %I2451.7 : Bool;
   "Carrier_42_SDCFaultCode" AT %IW2452 : Word;   // SDC FAULT CODE
   "Carrier_42_CarrierPosition" AT %ID2454 : DWord;   // CARRIER POSITION
   "Carrier_42_CarrierNumber" AT %IW2458 : Word;   // CARRIER NUMBER
   "Carrier_42_G120DControlWord" AT %IW2460 : Word;   // G120D_STW1_CONTROL
   "Carrier_42_G120DControlWord.0" AT %I2460.0 : Bool;   // Bit_00_ON
   "Carrier_42_G120DControlWord.1" AT %I2460.1 : Bool;   // Bit_01_AUS2_INH
   "Carrier_42_G120DControlWord.2" AT %I2460.2 : Bool;   // Bit_02_AUS3_STOP
   "Carrier_42_G120DControlWord.3" AT %I2460.3 : Bool;   // Bit_03_EN
